VERSION : 0.1
   VAR
      MC_Interface : Array[0..12] of Struct
         Data_from_MC : Struct   // Signal from the mould carrier to the machine
            Automatic_mode : Bool;   // Mouldcarrier is in automatic mode and ready for production
            Selected : Bool;   // Mouldcarrier is selected
            Shot_preperation : Bool;   // Set shot preperation
            Shot_release : Bool;   // Set shot release
            Robot_release : Bool;   // Release move robot into MC
            Vacuum_on : Bool;   // Vacuum pump on from MC
            CP_forward : Bool;   // Cleaning piston forward from MC
            Com_control : Bool;   // Communication control
            Toolcode : Byte;   // Toolcode from MC
            Temperature_1 : Int;   // Temperature 1 from MC
            Temperature_2 : Int;   // Temperature 2 from MC
            Angle_frame_foaming_pos : Real;   // Angle (°) frame in foaming position
            Spare_10 : Word;
            Spare_12 : Word;
            Spare_14 : Word;
         END_STRUCT;
         Data_to_MC : Struct   // Signal from the machine to the mould carrier
            Automatic_mode : Bool;   // Foaming machine ready for production
            Service_mode : Bool;   // Shot simmulation active
            MH_selected : Bool;   // Mixinghead is selected
            Shot_runs : Bool;   // Shot runs
            Shot_end : Bool;   // Shot end
            Fault : Bool;   // Fault during shot
            Robot_out_of_MC : Bool;   // Robot out of mould carrier (to close the MC)
            Com_Control : Bool;   // Communication control
            Toolcode : Byte;   // Toolcode copy from foaming machine
            Spare_2 : Word;
            Spare_4 : Word;
            Spare_6 : Word;
            Spare_8 : Word;
            Spare_10 : Word;
            Spare_12 : Word;
            Spare_14 : Word;
         END_STRUCT;
      END_STRUCT;
   END_VAR
BEGIN
   MC_Interface[0].Data_to_MC.Spare_8 := 16#0000;
   MC_Interface[0].Data_to_MC.Spare_6 := 16#0000;
   MC_Interface[0].Data_to_MC.Spare_4 := 16#0000;
   MC_Interface[0].Data_to_MC.Spare_2 := 16#0000;
   MC_Interface[0].Data_to_MC.Toolcode := 16#00;
   MC_Interface[0].Data_to_MC.Com_Control := FALSE;
   MC_Interface[0].Data_to_MC.Robot_out_of_MC := FALSE;
   MC_Interface[0].Data_to_MC.Fault := FALSE;
   MC_Interface[0].Data_to_MC.Shot_end := FALSE;
   MC_Interface[0].Data_to_MC.Shot_runs := FALSE;
   MC_Interface[0].Data_to_MC.MH_selected := FALSE;
   MC_Interface[0].Data_to_MC.Service_mode := FALSE;
   MC_Interface[0].Data_to_MC.Automatic_mode := FALSE;
   MC_Interface[0].Data_from_MC.Automatic_mode := FALSE;
   MC_Interface[0].Data_from_MC.Selected := FALSE;
   MC_Interface[0].Data_from_MC.Shot_preperation := FALSE;
   MC_Interface[0].Data_from_MC.Shot_release := FALSE;
   MC_Interface[0].Data_from_MC.Robot_release := FALSE;
   MC_Interface[0].Data_from_MC.Vacuum_on := FALSE;
   MC_Interface[0].Data_from_MC.CP_forward := FALSE;
   MC_Interface[0].Data_from_MC.Com_control := FALSE;
   MC_Interface[0].Data_from_MC.Toolcode := 16#02;
   MC_Interface[0].Data_from_MC.Temperature_1 := 16#0000;
   MC_Interface[0].Data_from_MC.Temperature_2 := 16#0000;
   MC_Interface[0].Data_from_MC.Angle_frame_foaming_pos := 16#0000;
END_DATA_BLOCK

DATA_BLOCK "DB009_Faults"   // DB9
TITLE = State signals of fault handling
{ S7_Optimized_Access := 'FALSE' }
AUTHOR : KT242
VERSION : 0.1
   VAR
      Fault_State_Grp_1_M1 : Bool := FALSE;   // In der Steuerung wurde eine Störung der Gruppe 1 der Maschine 1 festgestellt
      Fault_State_Grp_2_M1 : Bool := FALSE;   // In der Steuerung wurde eine Störung der Gruppe 2 der Maschine 1 festgestellt
      Fault_State_Grp_3_M1 : Bool := FALSE;   // In der Steuerung wurde eine Störung der Gruppe 3 der Maschine 1 festgestellt
      Fault_State_Grp_1_M2 : Bool := FALSE;   // In der Steuerung wurde eine Störung der Gruppe 1 der Maschine 2 festgestellt
      Fault_State_Grp_2_M2 : Bool := FALSE;   // In der Steuerung wurde eine Störung der Gruppe 2 der Maschine 2 festgestellt
      Fault_State_Grp_3_M2 : Bool := FALSE;   // In der Steuerung wurde eine Störung der Gruppe 3 der Maschine 2 festgestellt
      Fault_State_Grp_1_M3 : Bool := FALSE;   // In der Steuerung wurde eine Störung der Gruppe 1 der Maschine 3 festgestellt
      Fault_State_Grp_2_M3 : Bool := FALSE;   // In der Steuerung wurde eine Störung der Gruppe 2 der Maschine 3 festgestellt
      Fault_State_Grp_3_M3 : Bool := FALSE;   // In der Steuerung wurde eine Störung der Gruppe 3 der Maschine 3 festgestellt
      Fault_State_Grp_1_M4 : Bool := FALSE;   // In der Steuerung wurde eine Störung der Gruppe 1 der Maschine 4 festgestellt
      Fault_State_Grp_2_M4 : Bool := FALSE;   // In der Steuerung wurde eine Störung der Gruppe 2 der Maschine 4 festgestellt
      Fault_State_Grp_3_M4 : Bool := FALSE;   // In der Steuerung wurde eine Störung der Gruppe 3 der Maschine 4 festgestellt
      Fault_State_Grp_1_ExtP : Bool := FALSE;   // In der Steuerung wurde eine Störung der Gruppe 1 der Fremdanlage festgestellt
      Fault_State_Grp_2_ExtP : Bool := FALSE;   // In der Steuerung wurde eine Störung der Gruppe 2 der Fremdanlage festgestellt
      Fault_State_Grp_3_ExtP : Bool := FALSE;   // In der Steuerung wurde eine Störung der Gruppe 3 der Fremdanlage festgestellt
      Fault_State_Grp_1_3_Exist : Bool := FALSE;   // In der Steuerung wurde eine Störung der Gruppe 1- 3 festgestellt
      Faultschanging_M1 : Bool := FALSE;   // Änderungsbit für die Signalauswertung // Hupe+ Lampe Maschine 1
      Faultschanging_M2 : Bool := FALSE;   // Änderungsbit für die Signalauswertung // Hupe+ Lampe Maschine 2
      Faultschanging_M3 : Bool := FALSE;   // Änderungsbit für die Signalauswertung // Hupe+ Lampe Maschine 3
      Faultschanging_M4 : Bool := FALSE;   // Änderungsbit für die Signalauswertung // Hupe+ Lampe Maschine 4
      Faultschanging_ExtP : Bool := FALSE;   // Änderungsbit für die Signalauswertung // Hupe+ Lampe Fremdanlage
      Reserve_2_5 : Bool := FALSE;
      Reserve_2_6 : Bool := FALSE;
      Reserve_2_7 : Bool := FALSE;
      HF_FaultsQuitOB35 : Bool := FALSE;   // Resetbit for faults in OB 35
      HF_Faults_Quit : Bool := FALSE;   // Flankenhilfsmerker für die Störungsquittierung
      HF_Horn : Bool := FALSE;   // Hilfsmerker für die Hupenansteuerung
      Faults_Reset_FKT_M1 : Bool := FALSE;   // Störungsbildung in den Funktionen der Maschine 1 zurücksetzen
      Faults_Reset_FKT_M2 : Bool := FALSE;   // Störungsbildung in den Funktionen der Maschine 2 zurücksetzen
      Faults_Reset_FKT_M3 : Bool := FALSE;   // Störungsbildung in den Funktionen der Maschine 3 zurücksetzen
      Faults_Reset_FKT_M4 : Bool := FALSE;   // Störungsbildung in den Funktionen der Maschine 4 zurücksetzen
      Faults_Reset_FKT_ExtP : Bool := FALSE;   // Störungsbildung in den Funktionen der Fremdanlage zurücksetzen
      Faults_Reset_Group : Bool := FALSE;   // Störungsbildung in den Störungsbausteinenzurücksetzen
      FaultPC_Level_1 : Bool := FALSE;
      FaultPC_Level_2 : Bool := FALSE;
      FaultPC_Level_3 : Bool := FALSE;
      Spare_6_3 : Bool := FALSE;
      Spare_6_4 : Bool := FALSE;
      Faults_FKT_Grp_1_M1 : Bool := FALSE;   // In der Steuerung wurde eine Störung der Gruppe 1 der Maschine 1 festgestellt
      Faults_FKT_Grp_2_M1 : Bool := FALSE;   // In der Steuerung wurde eine Störung der Gruppe 2 der Maschine 1 festgestellt
      Faults_FKT_Grp_3_M1 : Bool := FALSE;   // In der Steuerung wurde eine Störung der Gruppe 3 der Maschine 1 festgestellt
      Faults_FKT_Grp_1_M2 : Bool := FALSE;   // In der Steuerung wurde eine Störung der Gruppe 1 der Maschine 2 festgestellt
      Faults_FKT_Grp_2_M2 : Bool := FALSE;   // In der Steuerung wurde eine Störung der Gruppe 2 der Maschine 2 festgestellt
      Faults_FKT_Grp_3_M2 : Bool := FALSE;   // In der Steuerung wurde eine Störung der Gruppe 3 der Maschine 2 festgestellt
      Faults_FKT_Grp_1_M3 : Bool := FALSE;   // In der Steuerung wurde eine Störung der Gruppe 1 der Maschine 3 festgestellt
      Faults_FKT_Grp_2_M3 : Bool := FALSE;   // In der Steuerung wurde eine Störung der Gruppe 2 der Maschine 3 festgestellt
      Faults_FKT_Grp_3_M3 : Bool := FALSE;   // In der Steuerung wurde eine Störung der Gruppe 3 der Maschine 3 festgestellt
      Faults_FKT_Grp_1_M4 : Bool := FALSE;   // In der Steuerung wurde eine Störung der Gruppe 1 der Maschine 4 festgestellt
      Faults_FKT_Grp_2_M4 : Bool := FALSE;   // In der Steuerung wurde eine Störung der Gruppe 2 der Maschine 4 festgestellt
      Faults_FKT_Grp_3_M4 : Bool := FALSE;   // In der Steuerung wurde eine Störung der Gruppe 3 der Maschine 4 festgestellt
      Faults_FKT_Grp_1_ExtP : Bool := FALSE;   // In der Steuerung wurde eine Störung der Gruppe 1 der Fremdanlage festgestellt
      Faults_FKT_Grp_2_ExtP : Bool := FALSE;   // In der Steuerung wurde eine Störung der Gruppe 2 der Fremdanlage festgestellt
      Faults_FKT_Grp_3_ExtP : Bool := FALSE;   // In der Steuerung wurde eine Störung der Gruppe 3 der Fremdanlage festgestellt
      Spare_8_7 : Bool := FALSE;
      NewMessage_M1 : Bool := FALSE;   // New message comes up at machine 1
      NewMessage_M2 : Bool := FALSE;   // New message comes up at machine 2
      NewMessage_M3 : Bool := FALSE;   // New message comes up at machine 3
      NewMessage_M4 : Bool := FALSE;   // New message comes up at machine 4
      GoneMessage_M1 : Bool := TRUE;   // Message is no longer active machine 1
      GoneMessage_M2 : Bool := FALSE;   // Message is no longer active machine 2
      GoneMessage_M3 : Bool := FALSE;   // Message is no longer active machine 3
      GoneMessage_M4 : Bool := FALSE;   // Message is no longer active machine 4
      MessageChangedToVisu : Bool := TRUE;   // Signal to visualisation -> show fault messages and messages
      MessageChangedNext : Bool := TRUE;
      Spare_10_02 : Bool := FALSE;
      Spare_10_03 : Bool := FALSE;
      Spare_10_04 : Bool := FALSE;
      Spare_10_05 : Bool := FALSE;
      Spare_10_06 : Bool := FALSE;
      Spare_10_07 : Bool := FALSE;
   END_VAR
BEGIN
END_DATA_BLOCK

DATA_BLOCK "DB_MouldEditor_HMI"   // DB10
{ S7_Optimized_Access := 'FALSE' }
VERSION : 0.1
   VAR
      uData : "typeMouldEditor_HMI";   // Data for mould editor HMI
   END_VAR
BEGIN
END_DATA_BLOCK

DATA_BLOCK "FB_MouldEditor_HMI_DB"   // DB13
{ S7_Optimized_Access := 'FALSE' }
VERSION : 0.1
"FB_MouldEditor_HMI"
BEGIN
END_DATA_BLOCK

DATA_BLOCK "DB14_TP_Shortcuts"   // DB14
{ S7_Optimized_Access := 'TRUE' }
VERSION : 0.1
   VAR
      TP_Shortcuts : Struct
         ButtonNo : Struct
            "0" : Bool := FALSE;
            "1" : Bool := FALSE;
            "2" : Bool := FALSE;
            "3" : Bool := FALSE;
            "4" : Bool := FALSE;
            "5" : Bool := FALSE;
            "6" : Bool := FALSE;
            "7" : Bool := FALSE;
         END_STRUCT;
         PageNo : Struct
            "0" : Int := 0;
            "1" : Int := 0;
            "2" : Int := 15;
            "3" : Int := 0;
            "4" : Int := 9;
            "5" : Int := 0;
            "6" : Int := 100;
            "7" : Int := 9020;
         END_STRUCT;
         Page_active : Struct
            "0" : Bool := FALSE;
            "1" : Bool := FALSE;
            "2" : Bool := FALSE;
            "3" : Bool := FALSE;
            "4" : Bool := FALSE;
            "5" : Bool := FALSE;
            "6" : Bool := FALSE;
            "7" : Bool := FALSE;
         END_STRUCT;
      END_STRUCT;
   END_VAR
BEGIN
END_DATA_BLOCK

DATA_BLOCK "DB025_Oszilloskop"   // DB25
{ S7_Optimized_Access := 'FALSE' }
VERSION : 0.1
   VAR
      Graph : Array[1..10] of Struct
         Auswahl : Int;
         Nummer : Int;
         Komponente : Int;
         Sensor : Int;
         DB_Nummer : Word;
         Adresse : Int;
         Skalierung : Real;
         Wert : Real;
         Bit : Int;
      END_STRUCT;
      SkalierungGraphLinks : Struct
         Startwert : Int := 0;
         Ebdwert : Int := 200;
      END_STRUCT;
      SkalierungGraphRechts : Struct
         Startwert : Int := 0;
         Ebdwert : Int := 220;
      END_STRUCT;
   END_VAR
BEGIN
   Graph[1].Skalierung := 1.0;
   Graph[2].Skalierung := 1.0;
   Graph[3].Skalierung := 1.0;
   Graph[4].Skalierung := 1.0;
   Graph[5].Skalierung := 1.0;
   Graph[6].Skalierung := 1.0;
   Graph[7].Skalierung := 1.0;
   Graph[8].Skalierung := 1.0;
   Graph[9].Skalierung := 1.0;
   Graph[10].Skalierung := 1.0;
   Graph[1].Auswahl := 30;
   Graph[1].Nummer := 0;
   Graph[1].Komponente := 1;
   Graph[1].Sensor := 1;
   Graph[1].DB_Nummer := 16#0000;
   Graph[1].Adresse := 0;
   Graph[1].Wert := 0.0;
   Graph[1].Bit := 0;
   Graph[2].Auswahl := 30;
   Graph[2].Nummer := 1;
   Graph[2].Komponente := 2;
   Graph[2].Sensor := 1;
   Graph[2].DB_Nummer := 16#0000;
   Graph[2].Adresse := 0;
   Graph[2].Wert := 0.0;
   Graph[2].Bit := 0;
   Graph[3].Auswahl := 0;
   Graph[3].Nummer := 0;
   Graph[3].Komponente := 0;
   Graph[3].Sensor := 0;
   Graph[3].DB_Nummer := 16#0000;
   Graph[3].Adresse := 0;
   Graph[3].Wert := 0.0;
   Graph[3].Bit := 0;
   Graph[4].Auswahl := 0;
   Graph[4].Nummer := 0;
   Graph[4].Komponente := 0;
   Graph[4].Sensor := 0;
   Graph[4].DB_Nummer := 16#0000;
   Graph[4].Adresse := 0;
   Graph[4].Wert := 0.0;
   Graph[4].Bit := 0;
   Graph[5].Auswahl := 0;
   Graph[5].Nummer := 0;
   Graph[5].Komponente := 0;
   Graph[5].Sensor := 0;
   Graph[5].DB_Nummer := 16#0000;
   Graph[5].Adresse := 0;
   Graph[5].Wert := 0.0;
   Graph[5].Bit := 0;
   Graph[6].Auswahl := 0;
   Graph[6].Nummer := 0;
   Graph[6].Komponente := 0;
   Graph[6].Sensor := 0;
   Graph[6].DB_Nummer := 16#0000;
   Graph[6].Adresse := 0;
   Graph[6].Wert := 0.0;
   Graph[6].Bit := 0;
   Graph[7].Auswahl := 20;
   Graph[7].Nummer := 1;
   Graph[7].Komponente := 1;
   Graph[7].Sensor := 2;
   Graph[7].DB_Nummer := 16#0000;
   Graph[7].Adresse := 0;
   Graph[7].Wert := 1.8;
   Graph[7].Bit := 0;
   Graph[8].Auswahl := 20;
   Graph[8].Nummer := 1;
   Graph[8].Komponente := 2;
   Graph[8].Sensor := 2;
   Graph[8].DB_Nummer := 16#0000;
   Graph[8].Adresse := 0;
   Graph[8].Wert := 2.2;
   Graph[8].Bit := 0;
   Graph[9].Auswahl := 0;
   Graph[9].Nummer := 0;
   Graph[9].Komponente := 0;
   Graph[9].Sensor := 0;
   Graph[9].DB_Nummer := 16#0000;
   Graph[9].Adresse := 0;
   Graph[9].Wert := 0.0;
   Graph[9].Bit := 0;
   Graph[10].Auswahl := 0;
   Graph[10].Nummer := 0;
   Graph[10].Komponente := 0;
   Graph[10].Sensor := 0;
   Graph[10].DB_Nummer := 16#0000;
   Graph[10].Adresse := 0;
   Graph[10].Wert := 0.0;
   Graph[10].Bit := 0;
END_DATA_BLOCK

DATA_BLOCK "BalluffReader_1"   // DB30
{ S7_Optimized_Access := 'FALSE' }
AUTHOR : Serrano
FAMILY : Ident
NAME : BIS60X2
VERSION : 1.8
"FB030_BallufReader"
BEGIN
END_DATA_BLOCK

DATA_BLOCK "BalluffReader_2"   // DB31
{ S7_Optimized_Access := 'FALSE' }
AUTHOR : Serrano
FAMILY : Ident
NAME : BIS60X2
VERSION : 1.8
"FB030_BallufReader"
BEGIN
END_DATA_BLOCK

DATA_BLOCK "BalluffReader"   // DB32
{ S7_Optimized_Access := 'FALSE' }
VERSION : 0.1
   VAR
      ReadWriteHead1 : Struct
         Command_Write : Bool := FALSE;
         FHM_Command_Write : Bool := FALSE;
         HM_Command_Write : Bool := FALSE;
         Command_Read : Bool := FALSE;
         FHM_Command_Read : Bool := FALSE;
         HM_Command_Read : Bool := FALSE;
         FHM_Read_Auto : Bool := FALSE;   // FHM Automatisch Lesen nach Schreiben
         HM_Read_Auto : Bool := FALSE;   // HM Automatisch Lesen nach Schreiben
         FHM_Code_was_readed : Bool := FALSE;   // FHM Code gelesen
         HM_Code_was_readed : Bool := FALSE;   // HM Code gelesen
         Code_was_readed : Bool := FALSE;   // HM Code gelesen
         FHM_Writing_was_activ : Bool := FALSE;   // FHM Beschreiben Datenträger war aktiv
         HM_Writing_was_activ : Bool := FALSE;   // HM Beschreiben Datenträger war aktiv
         FHM_Start_Zyklus : Bool;
         Spare_1_6 : Bool;
         Spare_1_7 : Bool;
         Fault_01 : Bool := FALSE;   // Kein Datenträger vorhanden
         Fault_02 : Bool := FALSE;   // Fehler beim Lesen
         Fault_03 : Bool := FALSE;   // Lesen abgebrochen, da Datenträger entfernt wurde
         Fault_04 : Bool := FALSE;   // Fehler beim Schreiben
         Fault_05 : Bool := FALSE;   // Schreiben abgebrochen, da Datenträger entfernt wurde
         Fault_06 : Bool := FALSE;   // Zugriffsfehler auf Speicher
         Fault_07 : Bool := FALSE;   // Falsche Befehlskennung oder Anzahl Byte bei einem Schreib-/Lesebefehl ist 0
         Fault_08 : Bool := FALSE;   // Kabelbruch des angewählten Schreib-/Lesekopfs
         Fault_09 : Bool := FALSE;   // EEProm in der Auswerteeinheit defekt
         Fault_10 : Bool := FALSE;   // Kommunikation zum Datenträger gestört
         Fault_11 : Bool := FALSE;   // Inhalt der 1. und 2. Bitleiste sind ungleich
         Fault_12 : Bool := FALSE;   // Startadresse + Anzahl Bytes > Speicherbereich in Initialisierung angegeben
         Fault_13 : Bool := FALSE;   // Ungültige max. Anzahl Schreibzyklen in Initialisierung angegeben
         Fault_14 : Bool := FALSE;   // max. Anzahl von 1kByte in Initialisierung überschritten
         Fault_15 : Bool := FALSE;   // Überwachung der Initialisierung bringt keine Übereinstimmung.
         Fault_16 : Bool := FALSE;   // Datenträger nicht initialisiert. Alle Bytes noch 00h
         Spare_4 : Byte;
         Spare_5 : Byte;
         Spare_6 : Byte;
         Spare_7 : Byte;
         TM_RFID : S5Time := S5T#4s;   // Überwachungszeit zum lesen/schreiben
         Send : Struct
            Program : Int;
            Text : Array[1..30] of Char;
         END_STRUCT;
         Receive : Struct
            Program : Int;
            Text : Array[1..30] of Char;
         END_STRUCT;
      END_STRUCT;
      ReadWriteHead2 : Struct
         Command_Write : Bool := FALSE;
         FHM_Command_Write : Bool := FALSE;
         HM_Command_Write : Bool := FALSE;
         Command_Read : Bool := FALSE;
         FHM_Command_Read : Bool := FALSE;
         HM_Command_Read : Bool := FALSE;
         FHM_Read_Auto : Bool := FALSE;   // FHM Automatisch Lesen nach Schreiben
         HM_Read_Auto : Bool := FALSE;   // HM Automatisch Lesen nach Schreiben
         FHM_Code_was_readed : Bool := FALSE;   // FHM Code gelesen
         HM_Code_was_readed : Bool := FALSE;   // HM Code gelesen
         Code_was_readed : Bool := FALSE;   // HM Code gelesen für Zylinder zurück
         FHM_Writing_was_activ : Bool := FALSE;   // FHM Beschreiben Datenträger war aktiv
         HM_Writing_was_activ : Bool := FALSE;   // HM Beschreiben Datenträger war aktiv
         FHM_Start_Zyklus : Bool;
         Spare_1_6 : Bool;
         Spare_1_7 : Bool;
         Fault_01 : Bool := FALSE;   // Kein Datenträger vorhanden
         Fault_02 : Bool := FALSE;   // Fehler beim Lesen
         Fault_03 : Bool := FALSE;   // Lesen abgebrochen, da Datenträger entfernt wurde
         Fault_04 : Bool := FALSE;   // Fehler beim Schreiben
         Fault_05 : Bool := FALSE;   // Schreiben abgebrochen, da Datenträger entfernt wurde
         Fault_06 : Bool := FALSE;   // Zugriffsfehler auf Speicher
         Fault_07 : Bool := FALSE;   // Falsche Befehlskennung oder Anzahl Byte bei einem Schreib-/Lesebefehl ist 0
         Fault_08 : Bool := FALSE;   // Kabelbruch des angewählten Schreib-/Lesekopfs
         Fault_09 : Bool := FALSE;   // EEProm in der Auswerteeinheit defekt
         Fault_10 : Bool := FALSE;   // Kommunikation zum Datenträger gestört
         Fault_11 : Bool := FALSE;   // Inhalt der 1. und 2. Bitleiste sind ungleich
         Fault_12 : Bool := FALSE;   // Startadresse + Anzahl Bytes > Speicherbereich in Initialisierung angegeben
         Fault_13 : Bool := FALSE;   // Ungültige max. Anzahl Schreibzyklen in Initialisierung angegeben
         Fault_14 : Bool := FALSE;   // max. Anzahl von 1kByte in Initialisierung überschritten
         Fault_15 : Bool := FALSE;   // Überwachung der Initialisierung bringt keine Übereinstimmung.
         Fault_16 : Bool := FALSE;   // Datenträger nicht initialisiert. Alle Bytes noch 00h
         Spare_4 : Byte;
         Spare_5 : Byte;
         Spare_6 : Byte;
         Spare_7 : Byte;
         TM_RFID : S5Time := S5T#4s;   // Überwachungszeit zum lesen/schreiben
         Send : Struct
            Program : Int;
            Text : Array[1..30] of Char;
         END_STRUCT;
         Receive : Struct
            Program : Int;
            Text : Array[1..30] of Char;
         END_STRUCT;
      END_STRUCT;
   END_VAR
BEGIN
END_DATA_BLOCK

DATA_BLOCK "DB110_Interf_Program_M1"   // DB110
TITLE = Signal between pouring machine and external plant parts
{ S7_Optimized_Access := 'FALSE' }
AUTHOR : KT242
VERSION : 0.1
   VAR
      Bits : Struct
         Ageflag : Bool := TRUE;
         Stop_Cycle : Bool := FALSE;
         startbutton_activated : Bool := FALSE;
         HF_StopCycleWHileToolDisabled : Bool := FALSE;
         F_StopCycleWHileToolDisabled : Bool := FALSE;
         LastShotAtThisMachine : Bool := FALSE;
         PulseShotEnd : Bool := FALSE;
         PulseToolFinished : Bool := FALSE;
         HF_FP_PulseToolFinished : Bool := TRUE;
         LockAutoCycleStart : Bool := FALSE;
         MouldNotReleased : Bool := FALSE;
         HF_FP_MouldNotReleased : Bool := FALSE;
         LastStandbyTimeTool : Bool := FALSE;
         PulseCycleEnd : Bool := FALSE;
         HF_FP_CycleNotRunning : Bool := TRUE;
         HF_FP_ResetProgramNo : Bool := FALSE;
      END_STRUCT;
      Putin_FIFOlist : "UDT001_DWord_1_32";
      FIRST : Int := 0;
      SECOND : Int := 0;
      FIFO : Struct
         FIFO_01 : Word := 16#0000;
         FIFO_02 : Word := 16#0000;
         FIFO_03 : Word := 16#0000;
         FIFO_04 : Word := 16#0000;
         FIFO_05 : Word := 16#0000;
         FIFO_06 : Word := 16#0000;
         FIFO_07 : Word := 16#0000;
         FIFO_08 : Word := 16#0000;
         FIFO_09 : Word := 16#0000;
         FIFO_10 : Word := 16#0000;
         FIFO_11 : Word := 16#0000;
         FIFO_12 : Word := 16#0000;
         FIFO_13 : Word := 16#0000;
         FIFO_14 : Word := 16#0000;
         FIFO_15 : Word := 16#0000;
         FIFO_16 : Word := 16#0000;
         FIFO_17 : Word := 16#0000;
         FIFO_18 : Word := 16#0000;
         FIFO_19 : Word := 16#0000;
         FIFO_20 : Word := 16#0000;
         FIFO_21 : Word := 16#0000;
         FIFO_22 : Word := 16#0000;
         FIFO_23 : Word := 16#0000;
         FIFO_24 : Word := 16#0000;
         FIFO_25 : Word := 16#0000;
         FIFO_26 : Word := 16#0000;
         FIFO_27 : Word := 16#0000;
         FIFO_28 : Word := 16#0000;
         FIFO_29 : Word := 16#0000;
         FIFO_30 : Word := 16#0000;
         FIFO_31 : Word := 16#0000;
         FIFO_32 : Word := 16#0000;
      END_STRUCT;
      Test_M01 : "UDT115_Test";
      Test_M02 : "UDT115_Test";
      Test_M03 : "UDT115_Test";
      Test_M04 : "UDT115_Test";
      Status_IF : Array[1..16] of "UDT112_IF_UP_MC";
      HM_MC_Fault : "UDT001_DWord_1_32";
      HM_MC_Shotend : "UDT001_DWord_1_32";
      HM_MC_Lamp : "UDT001_DWord_1_32";
      HM_MC_mould_Closing : "UDT001_DWord_1_32";
      HM_MC_spare : "UDT001_DWord_1_32";
      Program_is_active : "UDT001_DWord_1_32";
      Program_No_01 : Word := 16#0000;
      Program_No_02 : Word := 16#0000;
      Program_No_03 : Word := 16#0000;
      Program_No_04 : Word := 16#0000;
      Program_No_05 : Word := 16#0000;
      Program_No_06 : Word := 16#0000;
      Program_No_07 : Word := 16#0000;
      Program_No_08 : Word := 16#0000;
      Robot_01 : "ABB_IRC5_Status";
      Mixingheadcleaner_01 : "UDT118_MH_Cleaner";
      Bandfilter_01 : "UDT119_Bandfilter";
      Robot_02 : "ABB_IRC5_Status";
      Mixingheadcleaner_02 : "UDT118_MH_Cleaner";
      Bandfilter_02 : "UDT119_Bandfilter";
      MixingHeadNo : Int := 0;
      Signals_ExPlant : Array[1..4] of "UDT1114_IF_Signals";
      Status_ExPlant : Array[1..4] of "UDT114_IF_externalPlant";
   END_VAR
BEGIN
   Putin_FIFOlist."25" := FALSE;
   Putin_FIFOlist."26" := FALSE;
   Putin_FIFOlist."27" := FALSE;
   Putin_FIFOlist."28" := FALSE;
   Putin_FIFOlist."29" := FALSE;
   Putin_FIFOlist."30" := FALSE;
   Putin_FIFOlist."31" := FALSE;
   Putin_FIFOlist."32" := FALSE;
   Putin_FIFOlist."17" := FALSE;
   Putin_FIFOlist."18" := FALSE;
   Putin_FIFOlist."19" := FALSE;
   Putin_FIFOlist."20" := FALSE;
   Putin_FIFOlist."21" := FALSE;
   Putin_FIFOlist."22" := FALSE;
   Putin_FIFOlist."23" := FALSE;
   Putin_FIFOlist."24" := FALSE;
   Putin_FIFOlist."09" := FALSE;
   Putin_FIFOlist."10" := FALSE;
   Putin_FIFOlist."11" := FALSE;
   Putin_FIFOlist."12" := FALSE;
   Putin_FIFOlist."13" := FALSE;
   Putin_FIFOlist."14" := FALSE;
   Putin_FIFOlist."15" := FALSE;
   Putin_FIFOlist."16" := FALSE;
   Putin_FIFOlist."01" := FALSE;
   Putin_FIFOlist."02" := FALSE;
   Putin_FIFOlist."03" := FALSE;
   Putin_FIFOlist."04" := FALSE;
   Putin_FIFOlist."05" := FALSE;
   Putin_FIFOlist."06" := FALSE;
   Putin_FIFOlist."07" := FALSE;
   Putin_FIFOlist."08" := FALSE;
   Test_M01.Test_runs := FALSE;
   Test_M01.Test_K1 := FALSE;
   Test_M01.Test_K2 := FALSE;
   Test_M01.Test_K3 := FALSE;
   Test_M01.Test_K4 := FALSE;
   Test_M01.Start_to_Cycle := FALSE;
   Test_M01.Stop_to_Cycle := FALSE;
   Test_M01.Spare_0_7 := FALSE;
   Test_M01.Spare_Byte := 16#00;
   Test_M02.Test_runs := FALSE;
   Test_M02.Test_K1 := FALSE;
   Test_M02.Test_K2 := FALSE;
   Test_M02.Test_K3 := FALSE;
   Test_M02.Test_K4 := FALSE;
   Test_M02.Start_to_Cycle := FALSE;
   Test_M02.Stop_to_Cycle := FALSE;
   Test_M02.Spare_0_7 := FALSE;
   Test_M02.Spare_Byte := 16#00;
   Test_M03.Test_runs := FALSE;
   Test_M03.Test_K1 := FALSE;
   Test_M03.Test_K2 := FALSE;
   Test_M03.Test_K3 := FALSE;
   Test_M03.Test_K4 := FALSE;
   Test_M03.Start_to_Cycle := FALSE;
   Test_M03.Stop_to_Cycle := FALSE;
   Test_M03.Spare_0_7 := FALSE;
   Test_M03.Spare_Byte := 16#00;
   Test_M04.Test_runs := FALSE;
   Test_M04.Test_K1 := FALSE;
   Test_M04.Test_K2 := FALSE;
   Test_M04.Test_K3 := FALSE;
   Test_M04.Test_K4 := FALSE;
   Test_M04.Start_to_Cycle := FALSE;
   Test_M04.Stop_to_Cycle := FALSE;
   Test_M04.Spare_0_7 := FALSE;
   Test_M04.Spare_Byte := 16#00;
   HM_MC_Fault."25" := FALSE;
   HM_MC_Fault."26" := FALSE;
   HM_MC_Fault."27" := FALSE;
   HM_MC_Fault."28" := FALSE;
   HM_MC_Fault."29" := FALSE;
   HM_MC_Fault."30" := FALSE;
   HM_MC_Fault."31" := FALSE;
   HM_MC_Fault."32" := FALSE;
   HM_MC_Fault."17" := FALSE;
   HM_MC_Fault."18" := FALSE;
   HM_MC_Fault."19" := FALSE;
   HM_MC_Fault."20" := FALSE;
   HM_MC_Fault."21" := FALSE;
   HM_MC_Fault."22" := FALSE;
   HM_MC_Fault."23" := FALSE;
   HM_MC_Fault."24" := FALSE;
   HM_MC_Fault."09" := FALSE;
   HM_MC_Fault."10" := FALSE;
   HM_MC_Fault."11" := FALSE;
   HM_MC_Fault."12" := FALSE;
   HM_MC_Fault."13" := FALSE;
   HM_MC_Fault."14" := FALSE;
   HM_MC_Fault."15" := FALSE;
   HM_MC_Fault."16" := FALSE;
   HM_MC_Fault."01" := FALSE;
   HM_MC_Fault."02" := FALSE;
   HM_MC_Fault."03" := FALSE;
   HM_MC_Fault."04" := FALSE;
   HM_MC_Fault."05" := FALSE;
   HM_MC_Fault."06" := FALSE;
   HM_MC_Fault."07" := FALSE;
   HM_MC_Fault."08" := FALSE;
   HM_MC_Shotend."25" := FALSE;
   HM_MC_Shotend."26" := FALSE;
   HM_MC_Shotend."27" := FALSE;
   HM_MC_Shotend."28" := FALSE;
   HM_MC_Shotend."29" := FALSE;
   HM_MC_Shotend."30" := FALSE;
   HM_MC_Shotend."31" := FALSE;
   HM_MC_Shotend."32" := FALSE;
   HM_MC_Shotend."17" := FALSE;
   HM_MC_Shotend."18" := FALSE;
   HM_MC_Shotend."19" := FALSE;
   HM_MC_Shotend."20" := FALSE;
   HM_MC_Shotend."21" := FALSE;
   HM_MC_Shotend."22" := FALSE;
   HM_MC_Shotend."23" := FALSE;
   HM_MC_Shotend."24" := FALSE;
   HM_MC_Shotend."09" := FALSE;
   HM_MC_Shotend."10" := FALSE;
   HM_MC_Shotend."11" := FALSE;
   HM_MC_Shotend."12" := FALSE;
   HM_MC_Shotend."13" := FALSE;
   HM_MC_Shotend."14" := FALSE;
   HM_MC_Shotend."15" := FALSE;
   HM_MC_Shotend."16" := FALSE;
   HM_MC_Shotend."01" := FALSE;
   HM_MC_Shotend."02" := FALSE;
   HM_MC_Shotend."03" := FALSE;
   HM_MC_Shotend."04" := FALSE;
   HM_MC_Shotend."05" := FALSE;
   HM_MC_Shotend."06" := FALSE;
   HM_MC_Shotend."07" := FALSE;
   HM_MC_Shotend."08" := FALSE;
   HM_MC_Lamp."25" := FALSE;
   HM_MC_Lamp."26" := FALSE;
   HM_MC_Lamp."27" := FALSE;
   HM_MC_Lamp."28" := FALSE;
   HM_MC_Lamp."29" := FALSE;
   HM_MC_Lamp."30" := FALSE;
   HM_MC_Lamp."31" := FALSE;
   HM_MC_Lamp."32" := FALSE;
   HM_MC_Lamp."17" := FALSE;
   HM_MC_Lamp."18" := FALSE;
   HM_MC_Lamp."19" := FALSE;
   HM_MC_Lamp."20" := FALSE;
   HM_MC_Lamp."21" := FALSE;
   HM_MC_Lamp."22" := FALSE;
   HM_MC_Lamp."23" := FALSE;
   HM_MC_Lamp."24" := FALSE;
   HM_MC_Lamp."09" := FALSE;
   HM_MC_Lamp."10" := FALSE;
   HM_MC_Lamp."11" := FALSE;
   HM_MC_Lamp."12" := FALSE;
   HM_MC_Lamp."13" := FALSE;
   HM_MC_Lamp."14" := FALSE;
   HM_MC_Lamp."15" := FALSE;
   HM_MC_Lamp."16" := FALSE;
   HM_MC_Lamp."01" := FALSE;
   HM_MC_Lamp."02" := FALSE;
   HM_MC_Lamp."03" := FALSE;
   HM_MC_Lamp."04" := FALSE;
   HM_MC_Lamp."05" := FALSE;
   HM_MC_Lamp."06" := FALSE;
   HM_MC_Lamp."07" := FALSE;
   HM_MC_Lamp."08" := FALSE;
   HM_MC_mould_Closing."25" := FALSE;
   HM_MC_mould_Closing."26" := FALSE;
   HM_MC_mould_Closing."27" := FALSE;
   HM_MC_mould_Closing."28" := FALSE;
   HM_MC_mould_Closing."29" := FALSE;
   HM_MC_mould_Closing."30" := FALSE;
   HM_MC_mould_Closing."31" := FALSE;
   HM_MC_mould_Closing."32" := FALSE;
   HM_MC_mould_Closing."17" := FALSE;
   HM_MC_mould_Closing."18" := FALSE;
   HM_MC_mould_Closing."19" := FALSE;
   HM_MC_mould_Closing."20" := FALSE;
   HM_MC_mould_Closing."21" := FALSE;
   HM_MC_mould_Closing."22" := FALSE;
   HM_MC_mould_Closing."23" := FALSE;
   HM_MC_mould_Closing."24" := FALSE;
   HM_MC_mould_Closing."09" := FALSE;
   HM_MC_mould_Closing."10" := FALSE;
   HM_MC_mould_Closing."11" := FALSE;
   HM_MC_mould_Closing."12" := FALSE;
   HM_MC_mould_Closing."13" := FALSE;
   HM_MC_mould_Closing."14" := FALSE;
   HM_MC_mould_Closing."15" := FALSE;
   HM_MC_mould_Closing."16" := FALSE;
   HM_MC_mould_Closing."01" := FALSE;
   HM_MC_mould_Closing."02" := FALSE;
   HM_MC_mould_Closing."03" := FALSE;
   HM_MC_mould_Closing."04" := FALSE;
   HM_MC_mould_Closing."05" := FALSE;
   HM_MC_mould_Closing."06" := FALSE;
   HM_MC_mould_Closing."07" := FALSE;
   HM_MC_mould_Closing."08" := FALSE;
   HM_MC_spare."25" := FALSE;
   HM_MC_spare."26" := FALSE;
   HM_MC_spare."27" := FALSE;
   HM_MC_spare."28" := FALSE;
   // 962 more start values not shown
END_DATA_BLOCK

DATA_BLOCK "DB119_Interface_Visu"   // DB119
TITLE = Signal between pouring machine and external plant parts
{ S7_Optimized_Access := 'FALSE' }
AUTHOR : KT242
VERSION : 0.1
   VAR
      "Inv.PrgNr" : Bool := TRUE;
      Profibus : Bool := FALSE;
      Paritätsbit : Bool := FALSE;
      ReadWriteDeviceNo : Int := 0;
      CopyDeviceNO : Int := 0;
      Read : Bool := FALSE;
      Write : Bool := FALSE;
      Copy : Bool := FALSE;
      Activ : Bool := FALSE;
      MouldCarrer : Array[0..12] of "UDT1111_MouldCarrier";
      APInterface : Array[0..12] of "UDT1112_APInterface";
   END_VAR
BEGIN
   APInterface[0].PrgNo := 16#FF;
   APInterface[0].ExtP_OK := TRUE;
   APInterface[0].Strobe := TRUE;
   APInterface[0].StrobeInv := TRUE;
   APInterface[0].MH_open := TRUE;
   APInterface[0].CP_forward := TRUE;
   APInterface[0].Preparation := TRUE;
   APInterface[0].Start_Cleaning := TRUE;
   APInterface[0].Stop := TRUE;
   APInterface[0].PU_OK := TRUE;
   APInterface[0].Strobe_quitt := TRUE;
   APInterface[0].cycle_run := TRUE;
   APInterface[0].ready_for_shot := TRUE;
   APInterface[0].shot_run := TRUE;
   APInterface[0].shot_end := TRUE;
   APInterface[0].Service_mode := TRUE;
   APInterface[0].CP_is_forward := TRUE;
   APInterface[0].Cleaning_finished := TRUE;
   APInterface[0].Reserve31 := TRUE;
   MouldCarrer[0].Preparation := FALSE;
   MouldCarrer[0].StartFoaming := FALSE;
   MouldCarrer[0].IN_Spare_01 := FALSE;
   MouldCarrer[0].IN_Spare_02 := FALSE;
   MouldCarrer[0].IN_Spare_03 := FALSE;
   MouldCarrer[0].IN_Spare_04 := FALSE;
   MouldCarrer[0].IN_Spare_05 := FALSE;
   MouldCarrer[0].IN_Spare_06 := FALSE;
   MouldCarrer[0].ShotEnds := FALSE;
   MouldCarrer[0].Break := FALSE;
   MouldCarrer[0].OUT_Spare_01 := FALSE;
   MouldCarrer[0].OUT_Spare_02 := FALSE;
   MouldCarrer[0].OUT_Spare_03 := FALSE;
   MouldCarrer[0].OUT_Spare_04 := FALSE;
   MouldCarrer[0].OUT_Spare_05 := FALSE;
   MouldCarrer[0].OUT_Spare_06 := FALSE;
   MouldCarrer[0].NoFault := FALSE;
   MouldCarrer[0].MachineAutomatic := FALSE;
   MouldCarrer[0].MHAutomatic := FALSE;
   MouldCarrer[0].RobotAutomatic := FALSE;
   MouldCarrer[0].WetShot := FALSE;
   MouldCarrer[0].CycleRun := FALSE;
   MouldCarrer[0].ReadyForShot := FALSE;
   MouldCarrer[0].ShotRun := FALSE;
   MouldCarrer[0].CPsisForward := FALSE;
   MouldCarrer[0].Status_Spare_01 := FALSE;
   MouldCarrer[0].Status_Spare_02 := FALSE;
   MouldCarrer[0].Status_Spare_03 := FALSE;
   MouldCarrer[0].Status_Spare_04 := FALSE;
   MouldCarrer[0].Status_Spare_05 := FALSE;
   MouldCarrer[0].Status_Spare_06 := FALSE;
   MouldCarrer[0].Status_Spare_07 := FALSE;
   MouldCarrer[0].ProgNumber := FALSE;
   MouldCarrer[0].Fault_01 := FALSE;
   MouldCarrer[0].Fault_02 := FALSE;
   MouldCarrer[0].Fault_03 := FALSE;
   MouldCarrer[0].Fault_04 := FALSE;
   MouldCarrer[0].Fault_05 := FALSE;
   MouldCarrer[0].Fault_06 := FALSE;
   MouldCarrer[0].Fault_07 := FALSE;
   MouldCarrer[0].Fault_08 := FALSE;
   MouldCarrer[1].Preparation := FALSE;
   MouldCarrer[1].StartFoaming := FALSE;
   MouldCarrer[1].IN_Spare_01 := FALSE;
   MouldCarrer[1].IN_Spare_02 := FALSE;
   MouldCarrer[1].IN_Spare_03 := FALSE;
   MouldCarrer[1].IN_Spare_04 := FALSE;
   MouldCarrer[1].IN_Spare_05 := FALSE;
   MouldCarrer[1].IN_Spare_06 := FALSE;
   MouldCarrer[1].ShotEnds := FALSE;
   MouldCarrer[1].Break := FALSE;
   MouldCarrer[1].OUT_Spare_01 := FALSE;
   MouldCarrer[1].OUT_Spare_02 := FALSE;
   MouldCarrer[1].OUT_Spare_03 := FALSE;
   MouldCarrer[1].OUT_Spare_04 := FALSE;
   MouldCarrer[1].OUT_Spare_05 := FALSE;
   MouldCarrer[1].OUT_Spare_06 := FALSE;
   MouldCarrer[1].NoFault := FALSE;
   MouldCarrer[1].MachineAutomatic := FALSE;
   MouldCarrer[1].MHAutomatic := FALSE;
   MouldCarrer[1].RobotAutomatic := FALSE;
   MouldCarrer[1].WetShot := FALSE;
   MouldCarrer[1].CycleRun := FALSE;
   MouldCarrer[1].ReadyForShot := FALSE;
   MouldCarrer[1].ShotRun := FALSE;
   MouldCarrer[1].CPsisForward := FALSE;
   MouldCarrer[1].Status_Spare_01 := FALSE;
   MouldCarrer[1].Status_Spare_02 := FALSE;
   MouldCarrer[1].Status_Spare_03 := FALSE;
   MouldCarrer[1].Status_Spare_04 := FALSE;
   MouldCarrer[1].Status_Spare_05 := FALSE;
   MouldCarrer[1].Status_Spare_06 := FALSE;
   MouldCarrer[1].Status_Spare_07 := FALSE;
   MouldCarrer[1].ProgNumber := FALSE;
   MouldCarrer[1].Fault_01 := FALSE;
   MouldCarrer[1].Fault_02 := FALSE;
   MouldCarrer[1].Fault_03 := FALSE;
   MouldCarrer[1].Fault_04 := FALSE;
   MouldCarrer[1].Fault_05 := FALSE;
   MouldCarrer[1].Fault_06 := FALSE;
   MouldCarrer[1].Fault_07 := FALSE;
   MouldCarrer[1].Fault_08 := FALSE;
   MouldCarrer[2].Preparation := FALSE;
   MouldCarrer[2].StartFoaming := FALSE;
   MouldCarrer[2].IN_Spare_01 := FALSE;
   MouldCarrer[2].IN_Spare_02 := FALSE;
   MouldCarrer[2].IN_Spare_03 := FALSE;
   MouldCarrer[2].IN_Spare_04 := FALSE;
   MouldCarrer[2].IN_Spare_05 := FALSE;
   MouldCarrer[2].IN_Spare_06 := FALSE;
   MouldCarrer[2].ShotEnds := FALSE;
   MouldCarrer[2].Break := FALSE;
   MouldCarrer[2].OUT_Spare_01 := FALSE;
   MouldCarrer[2].OUT_Spare_02 := FALSE;
   MouldCarrer[2].OUT_Spare_03 := FALSE;
   MouldCarrer[2].OUT_Spare_04 := FALSE;
   MouldCarrer[2].OUT_Spare_05 := FALSE;
   MouldCarrer[2].OUT_Spare_06 := FALSE;
   MouldCarrer[2].NoFault := FALSE;
   MouldCarrer[2].MachineAutomatic := FALSE;
   MouldCarrer[2].MHAutomatic := FALSE;
   MouldCarrer[2].RobotAutomatic := FALSE;
   MouldCarrer[2].WetShot := FALSE;
   MouldCarrer[2].CycleRun := FALSE;
   MouldCarrer[2].ReadyForShot := FALSE;
   MouldCarrer[2].ShotRun := FALSE;
   MouldCarrer[2].CPsisForward := FALSE;
   MouldCarrer[2].Status_Spare_01 := FALSE;
   MouldCarrer[2].Status_Spare_02 := FALSE;
   MouldCarrer[2].Status_Spare_03 := FALSE;
   MouldCarrer[2].Status_Spare_04 := FALSE;
   MouldCarrer[2].Status_Spare_05 := FALSE;
   MouldCarrer[2].Status_Spare_06 := FALSE;
   MouldCarrer[2].Status_Spare_07 := FALSE;
   MouldCarrer[2].ProgNumber := FALSE;
   MouldCarrer[2].Fault_01 := FALSE;
   MouldCarrer[2].Fault_02 := FALSE;
   MouldCarrer[2].Fault_03 := FALSE;
   MouldCarrer[2].Fault_04 := FALSE;
   MouldCarrer[2].Fault_05 := FALSE;
   MouldCarrer[2].Fault_06 := FALSE;
   MouldCarrer[2].Fault_07 := FALSE;
   MouldCarrer[2].Fault_08 := FALSE;
   MouldCarrer[3].Preparation := FALSE;
   MouldCarrer[3].StartFoaming := FALSE;
   MouldCarrer[3].IN_Spare_01 := FALSE;
   MouldCarrer[3].IN_Spare_02 := FALSE;
   MouldCarrer[3].IN_Spare_03 := FALSE;
   MouldCarrer[3].IN_Spare_04 := FALSE;
   MouldCarrer[3].IN_Spare_05 := FALSE;
   MouldCarrer[3].IN_Spare_06 := FALSE;
   MouldCarrer[3].ShotEnds := FALSE;
   MouldCarrer[3].Break := FALSE;
   MouldCarrer[3].OUT_Spare_01 := FALSE;
   MouldCarrer[3].OUT_Spare_02 := FALSE;
   MouldCarrer[3].OUT_Spare_03 := FALSE;
   MouldCarrer[3].OUT_Spare_04 := FALSE;
   MouldCarrer[3].OUT_Spare_05 := FALSE;
   MouldCarrer[3].OUT_Spare_06 := FALSE;
   MouldCarrer[3].NoFault := FALSE;
   MouldCarrer[3].MachineAutomatic := FALSE;
   MouldCarrer[3].MHAutomatic := FALSE;
   MouldCarrer[3].RobotAutomatic := FALSE;
   MouldCarrer[3].WetShot := FALSE;
   MouldCarrer[3].CycleRun := FALSE;
   MouldCarrer[3].ReadyForShot := FALSE;
   MouldCarrer[3].ShotRun := FALSE;
   MouldCarrer[3].CPsisForward := FALSE;
   MouldCarrer[3].Status_Spare_01 := FALSE;
   MouldCarrer[3].Status_Spare_02 := FALSE;
   MouldCarrer[3].Status_Spare_03 := FALSE;
   MouldCarrer[3].Status_Spare_04 := FALSE;
   MouldCarrer[3].Status_Spare_05 := FALSE;
   MouldCarrer[3].Status_Spare_06 := FALSE;
   MouldCarrer[3].Status_Spare_07 := FALSE;
   MouldCarrer[3].ProgNumber := FALSE;
   MouldCarrer[3].Fault_01 := FALSE;
   MouldCarrer[3].Fault_02 := FALSE;
   MouldCarrer[3].Fault_03 := FALSE;
   MouldCarrer[3].Fault_04 := FALSE;
   MouldCarrer[3].Fault_05 := FALSE;
   MouldCarrer[3].Fault_06 := FALSE;
   MouldCarrer[3].Fault_07 := FALSE;
   MouldCarrer[3].Fault_08 := FALSE;
   MouldCarrer[4].Preparation := FALSE;
   MouldCarrer[4].StartFoaming := FALSE;
   MouldCarrer[4].IN_Spare_01 := FALSE;
   MouldCarrer[4].IN_Spare_02 := FALSE;
   MouldCarrer[4].IN_Spare_03 := FALSE;
   MouldCarrer[4].IN_Spare_04 := FALSE;
   MouldCarrer[4].IN_Spare_05 := FALSE;
   MouldCarrer[4].IN_Spare_06 := FALSE;
   MouldCarrer[4].ShotEnds := FALSE;
   MouldCarrer[4].Break := FALSE;
   MouldCarrer[4].OUT_Spare_01 := FALSE;
   MouldCarrer[4].OUT_Spare_02 := FALSE;
   MouldCarrer[4].OUT_Spare_03 := FALSE;
   MouldCarrer[4].OUT_Spare_04 := FALSE;
   MouldCarrer[4].OUT_Spare_05 := FALSE;
   MouldCarrer[4].OUT_Spare_06 := FALSE;
   MouldCarrer[4].NoFault := FALSE;
   // 983 more start values not shown
END_DATA_BLOCK

DATA_BLOCK "DB122_FlowIndexState"   // DB122
TITLE = Flow-Index and Flow-State of modul-channel
{ S7_Optimized_Access := 'FALSE' }
AUTHOR : KT242
NAME : Flow
VERSION : 0.1
   VAR
      MeteringUnit : Array[0..12] of "UDT121_DF_Chanel";
   END_VAR
BEGIN
   MeteringUnit[0].OUT_PROCAN.FlowIndex.FlowIndex0 := FALSE;
   MeteringUnit[0].OUT_PROCAN.FlowIndex.FlowIndex1 := FALSE;
   MeteringUnit[0].OUT_PROCAN.FlowIndex.FlowIndex2 := FALSE;
   MeteringUnit[0].OUT_PROCAN.FlowIndex.FlowIndex3 := FALSE;
   MeteringUnit[0].OUT_PROCAN.FlowIndex.Spare4 := FALSE;
   MeteringUnit[0].OUT_PROCAN.FlowIndex.Notclosedloop := FALSE;
   MeteringUnit[0].OUT_PROCAN.FlowIndex.StartQPB := FALSE;
   MeteringUnit[0].OUT_PROCAN.FlowIndex.Enableclosedloop := FALSE;
   MeteringUnit[0].OUT_PROCAN.TandemComand := 16#0000;
   MeteringUnit[0].OUT_PROCAN.SpareWord := 16#0000;
   MeteringUnit[0].OUT_PROCAN.Spare_DWORD_56 := 16#0000_0000;
   MeteringUnit[0].IN_PROCAN.Flowrate := 0;
   MeteringUnit[0].IN_PROCAN.PistonPosition := 0;
   MeteringUnit[0].IN_PROCAN.TandemStatus := 16#0000;
   MeteringUnit[0].IN_PROCAN.Spare_DWORD_96 := 16#0000_0000;
   MeteringUnit[1].OUT_PROCAN.FlowIndex.FlowIndex0 := FALSE;
   MeteringUnit[1].OUT_PROCAN.FlowIndex.FlowIndex1 := FALSE;
   MeteringUnit[1].OUT_PROCAN.FlowIndex.FlowIndex2 := FALSE;
   MeteringUnit[1].OUT_PROCAN.FlowIndex.FlowIndex3 := FALSE;
   MeteringUnit[1].OUT_PROCAN.FlowIndex.Spare4 := FALSE;
   MeteringUnit[1].OUT_PROCAN.FlowIndex.Notclosedloop := FALSE;
   MeteringUnit[1].OUT_PROCAN.FlowIndex.StartQPB := FALSE;
   MeteringUnit[1].OUT_PROCAN.FlowIndex.Enableclosedloop := FALSE;
   MeteringUnit[1].OUT_PROCAN.TandemComand := 16#0000;
   MeteringUnit[1].OUT_PROCAN.SpareWord := 16#0000;
   MeteringUnit[1].OUT_PROCAN.Spare_DWORD_56 := 16#0000_0000;
   MeteringUnit[1].IN_PROCAN.Flowrate := 0;
   MeteringUnit[1].IN_PROCAN.PistonPosition := 0;
   MeteringUnit[1].IN_PROCAN.TandemStatus := 16#0000;
   MeteringUnit[1].IN_PROCAN.Spare_DWORD_96 := 16#0000_0000;
   MeteringUnit[2].OUT_PROCAN.FlowIndex.FlowIndex0 := FALSE;
   MeteringUnit[2].OUT_PROCAN.FlowIndex.FlowIndex1 := FALSE;
   MeteringUnit[2].OUT_PROCAN.FlowIndex.FlowIndex2 := FALSE;
   MeteringUnit[2].OUT_PROCAN.FlowIndex.FlowIndex3 := FALSE;
   MeteringUnit[2].OUT_PROCAN.FlowIndex.Spare4 := FALSE;
   MeteringUnit[2].OUT_PROCAN.FlowIndex.Notclosedloop := FALSE;
   MeteringUnit[2].OUT_PROCAN.FlowIndex.StartQPB := FALSE;
   MeteringUnit[2].OUT_PROCAN.FlowIndex.Enableclosedloop := FALSE;
   MeteringUnit[2].OUT_PROCAN.TandemComand := 16#0000;
   MeteringUnit[2].OUT_PROCAN.SpareWord := 16#0000;
   MeteringUnit[2].OUT_PROCAN.Spare_DWORD_56 := 16#0000_0000;
   MeteringUnit[2].IN_PROCAN.Flowrate := 0;
   MeteringUnit[2].IN_PROCAN.PistonPosition := 0;
   MeteringUnit[2].IN_PROCAN.TandemStatus := 16#0000;
   MeteringUnit[2].IN_PROCAN.Spare_DWORD_96 := 16#0000_0000;
   MeteringUnit[3].OUT_PROCAN.FlowIndex.FlowIndex0 := FALSE;
   MeteringUnit[3].OUT_PROCAN.FlowIndex.FlowIndex1 := FALSE;
   MeteringUnit[3].OUT_PROCAN.FlowIndex.FlowIndex2 := FALSE;
   MeteringUnit[3].OUT_PROCAN.FlowIndex.FlowIndex3 := FALSE;
   MeteringUnit[3].OUT_PROCAN.FlowIndex.Spare4 := FALSE;
   MeteringUnit[3].OUT_PROCAN.FlowIndex.Notclosedloop := FALSE;
   MeteringUnit[3].OUT_PROCAN.FlowIndex.StartQPB := FALSE;
   MeteringUnit[3].OUT_PROCAN.FlowIndex.Enableclosedloop := FALSE;
   MeteringUnit[3].OUT_PROCAN.TandemComand := 16#0000;
   MeteringUnit[3].OUT_PROCAN.SpareWord := 16#0000;
   MeteringUnit[3].OUT_PROCAN.Spare_DWORD_56 := 16#0000_0000;
   MeteringUnit[3].IN_PROCAN.Flowrate := 0;
   MeteringUnit[3].IN_PROCAN.PistonPosition := 0;
   MeteringUnit[3].IN_PROCAN.TandemStatus := 16#0000;
   MeteringUnit[3].IN_PROCAN.Spare_DWORD_96 := 16#0000_0000;
   MeteringUnit[4].OUT_PROCAN.FlowIndex.FlowIndex0 := FALSE;
   MeteringUnit[4].OUT_PROCAN.FlowIndex.FlowIndex1 := FALSE;
   MeteringUnit[4].OUT_PROCAN.FlowIndex.FlowIndex2 := FALSE;
   MeteringUnit[4].OUT_PROCAN.FlowIndex.FlowIndex3 := FALSE;
   MeteringUnit[4].OUT_PROCAN.FlowIndex.Spare4 := FALSE;
   MeteringUnit[4].OUT_PROCAN.FlowIndex.Notclosedloop := FALSE;
   MeteringUnit[4].OUT_PROCAN.FlowIndex.StartQPB := FALSE;
   MeteringUnit[4].OUT_PROCAN.FlowIndex.Enableclosedloop := FALSE;
   MeteringUnit[4].OUT_PROCAN.TandemComand := 16#0000;
   MeteringUnit[4].OUT_PROCAN.SpareWord := 16#0000;
   MeteringUnit[4].OUT_PROCAN.Spare_DWORD_56 := 16#0000_0000;
   MeteringUnit[4].IN_PROCAN.Flowrate := 0;
   MeteringUnit[4].IN_PROCAN.PistonPosition := 0;
   MeteringUnit[4].IN_PROCAN.TandemStatus := 16#0000;
   MeteringUnit[4].IN_PROCAN.Spare_DWORD_96 := 16#0000_0000;
   MeteringUnit[5].OUT_PROCAN.FlowIndex.FlowIndex0 := FALSE;
   MeteringUnit[5].OUT_PROCAN.FlowIndex.FlowIndex1 := FALSE;
   MeteringUnit[5].OUT_PROCAN.FlowIndex.FlowIndex2 := FALSE;
   MeteringUnit[5].OUT_PROCAN.FlowIndex.FlowIndex3 := FALSE;
   MeteringUnit[5].OUT_PROCAN.FlowIndex.Spare4 := FALSE;
   MeteringUnit[5].OUT_PROCAN.FlowIndex.Notclosedloop := FALSE;
   MeteringUnit[5].OUT_PROCAN.FlowIndex.StartQPB := FALSE;
   MeteringUnit[5].OUT_PROCAN.FlowIndex.Enableclosedloop := FALSE;
   MeteringUnit[5].OUT_PROCAN.TandemComand := 16#0000;
   MeteringUnit[5].OUT_PROCAN.SpareWord := 16#0000;
   MeteringUnit[5].OUT_PROCAN.Spare_DWORD_56 := 16#0000_0000;
   MeteringUnit[5].IN_PROCAN.Flowrate := 0;
   MeteringUnit[5].IN_PROCAN.PistonPosition := 0;
   MeteringUnit[5].IN_PROCAN.TandemStatus := 16#0000;
   MeteringUnit[5].IN_PROCAN.Spare_DWORD_96 := 16#0000_0000;
   MeteringUnit[6].OUT_PROCAN.FlowIndex.FlowIndex0 := FALSE;
   MeteringUnit[6].OUT_PROCAN.FlowIndex.FlowIndex1 := FALSE;
   MeteringUnit[6].OUT_PROCAN.FlowIndex.FlowIndex2 := FALSE;
   MeteringUnit[6].OUT_PROCAN.FlowIndex.FlowIndex3 := FALSE;
   MeteringUnit[6].OUT_PROCAN.FlowIndex.Spare4 := FALSE;
   MeteringUnit[6].OUT_PROCAN.FlowIndex.Notclosedloop := FALSE;
   MeteringUnit[6].OUT_PROCAN.FlowIndex.StartQPB := FALSE;
   MeteringUnit[6].OUT_PROCAN.FlowIndex.Enableclosedloop := FALSE;
   MeteringUnit[6].OUT_PROCAN.TandemComand := 16#0000;
   MeteringUnit[6].OUT_PROCAN.SpareWord := 16#0000;
   MeteringUnit[6].OUT_PROCAN.Spare_DWORD_56 := 16#0000_0000;
   MeteringUnit[6].IN_PROCAN.Flowrate := 0;
   MeteringUnit[6].IN_PROCAN.PistonPosition := 0;
   MeteringUnit[6].IN_PROCAN.TandemStatus := 16#0000;
   MeteringUnit[6].IN_PROCAN.Spare_DWORD_96 := 16#0000_0000;
   MeteringUnit[7].OUT_PROCAN.FlowIndex.FlowIndex0 := FALSE;
   MeteringUnit[7].OUT_PROCAN.FlowIndex.FlowIndex1 := FALSE;
   MeteringUnit[7].OUT_PROCAN.FlowIndex.FlowIndex2 := FALSE;
   MeteringUnit[7].OUT_PROCAN.FlowIndex.FlowIndex3 := FALSE;
   MeteringUnit[7].OUT_PROCAN.FlowIndex.Spare4 := FALSE;
   MeteringUnit[7].OUT_PROCAN.FlowIndex.Notclosedloop := FALSE;
   MeteringUnit[7].OUT_PROCAN.FlowIndex.StartQPB := FALSE;
   MeteringUnit[7].OUT_PROCAN.FlowIndex.Enableclosedloop := FALSE;
   MeteringUnit[7].OUT_PROCAN.TandemComand := 16#0000;
   MeteringUnit[7].OUT_PROCAN.SpareWord := 16#0000;
   MeteringUnit[7].OUT_PROCAN.Spare_DWORD_56 := 16#0000_0000;
   MeteringUnit[7].IN_PROCAN.Flowrate := 0;
   MeteringUnit[7].IN_PROCAN.PistonPosition := 0;
   MeteringUnit[7].IN_PROCAN.TandemStatus := 16#0000;
   MeteringUnit[7].IN_PROCAN.Spare_DWORD_96 := 16#0000_0000;
   MeteringUnit[8].OUT_PROCAN.FlowIndex.FlowIndex0 := FALSE;
   MeteringUnit[8].OUT_PROCAN.FlowIndex.FlowIndex1 := FALSE;
   MeteringUnit[8].OUT_PROCAN.FlowIndex.FlowIndex2 := FALSE;
   MeteringUnit[8].OUT_PROCAN.FlowIndex.FlowIndex3 := FALSE;
   MeteringUnit[8].OUT_PROCAN.FlowIndex.Spare4 := FALSE;
   MeteringUnit[8].OUT_PROCAN.FlowIndex.Notclosedloop := FALSE;
   MeteringUnit[8].OUT_PROCAN.FlowIndex.StartQPB := FALSE;
   MeteringUnit[8].OUT_PROCAN.FlowIndex.Enableclosedloop := FALSE;
   MeteringUnit[8].OUT_PROCAN.TandemComand := 16#0000;
   MeteringUnit[8].OUT_PROCAN.SpareWord := 16#0000;
   MeteringUnit[8].OUT_PROCAN.Spare_DWORD_56 := 16#0000_0000;
   MeteringUnit[8].IN_PROCAN.Flowrate := 0;
   MeteringUnit[8].IN_PROCAN.PistonPosition := 0;
   MeteringUnit[8].IN_PROCAN.TandemStatus := 16#0000;
   MeteringUnit[8].IN_PROCAN.Spare_DWORD_96 := 16#0000_0000;
   MeteringUnit[9].OUT_PROCAN.FlowIndex.FlowIndex0 := FALSE;
   MeteringUnit[9].OUT_PROCAN.FlowIndex.FlowIndex1 := FALSE;
   MeteringUnit[9].OUT_PROCAN.FlowIndex.FlowIndex2 := FALSE;
   MeteringUnit[9].OUT_PROCAN.FlowIndex.FlowIndex3 := FALSE;
   MeteringUnit[9].OUT_PROCAN.FlowIndex.Spare4 := FALSE;
   MeteringUnit[9].OUT_PROCAN.FlowIndex.Notclosedloop := FALSE;
   MeteringUnit[9].OUT_PROCAN.FlowIndex.StartQPB := FALSE;
   MeteringUnit[9].OUT_PROCAN.FlowIndex.Enableclosedloop := FALSE;
   MeteringUnit[9].OUT_PROCAN.TandemComand := 16#0000;
   MeteringUnit[9].OUT_PROCAN.SpareWord := 16#0000;
   MeteringUnit[9].OUT_PROCAN.Spare_DWORD_56 := 16#0000_0000;
   MeteringUnit[9].IN_PROCAN.Flowrate := 0;
   MeteringUnit[9].IN_PROCAN.PistonPosition := 0;
   MeteringUnit[9].IN_PROCAN.TandemStatus := 16#0000;
   MeteringUnit[9].IN_PROCAN.Spare_DWORD_96 := 16#0000_0000;
   MeteringUnit[10].OUT_PROCAN.FlowIndex.FlowIndex0 := FALSE;
   MeteringUnit[10].OUT_PROCAN.FlowIndex.FlowIndex1 := FALSE;
   MeteringUnit[10].OUT_PROCAN.FlowIndex.FlowIndex2 := FALSE;
   MeteringUnit[10].OUT_PROCAN.FlowIndex.FlowIndex3 := FALSE;
   MeteringUnit[10].OUT_PROCAN.FlowIndex.Spare4 := FALSE;
   MeteringUnit[10].OUT_PROCAN.FlowIndex.Notclosedloop := FALSE;
   MeteringUnit[10].OUT_PROCAN.FlowIndex.StartQPB := FALSE;
   MeteringUnit[10].OUT_PROCAN.FlowIndex.Enableclosedloop := FALSE;
   MeteringUnit[10].OUT_PROCAN.TandemComand := 16#0000;
   MeteringUnit[10].OUT_PROCAN.SpareWord := 16#0000;
   MeteringUnit[10].OUT_PROCAN.Spare_DWORD_56 := 16#0000_0000;
   MeteringUnit[10].IN_PROCAN.Flowrate := 0;
   MeteringUnit[10].IN_PROCAN.PistonPosition := 0;
   MeteringUnit[10].IN_PROCAN.TandemStatus := 16#0000;
   MeteringUnit[10].IN_PROCAN.Spare_DWORD_96 := 16#0000_0000;
   MeteringUnit[11].OUT_PROCAN.FlowIndex.FlowIndex0 := FALSE;
   MeteringUnit[11].OUT_PROCAN.FlowIndex.FlowIndex1 := FALSE;
   MeteringUnit[11].OUT_PROCAN.FlowIndex.FlowIndex2 := FALSE;
   MeteringUnit[11].OUT_PROCAN.FlowIndex.FlowIndex3 := FALSE;
   MeteringUnit[11].OUT_PROCAN.FlowIndex.Spare4 := FALSE;
   MeteringUnit[11].OUT_PROCAN.FlowIndex.Notclosedloop := FALSE;
   MeteringUnit[11].OUT_PROCAN.FlowIndex.StartQPB := FALSE;
   MeteringUnit[11].OUT_PROCAN.FlowIndex.Enableclosedloop := FALSE;
   MeteringUnit[11].OUT_PROCAN.TandemComand := 16#0000;
   MeteringUnit[11].OUT_PROCAN.SpareWord := 16#0000;
   MeteringUnit[11].OUT_PROCAN.Spare_DWORD_56 := 16#0000_0000;
   MeteringUnit[11].IN_PROCAN.Flowrate := 0;
   MeteringUnit[11].IN_PROCAN.PistonPosition := 0;
   MeteringUnit[11].IN_PROCAN.TandemStatus := 16#0000;
   MeteringUnit[11].IN_PROCAN.Spare_DWORD_96 := 16#0000_0000;
   MeteringUnit[12].OUT_PROCAN.FlowIndex.FlowIndex0 := FALSE;
   MeteringUnit[12].OUT_PROCAN.FlowIndex.FlowIndex1 := FALSE;
   MeteringUnit[12].OUT_PROCAN.FlowIndex.FlowIndex2 := FALSE;
   MeteringUnit[12].OUT_PROCAN.FlowIndex.FlowIndex3 := FALSE;
   MeteringUnit[12].OUT_PROCAN.FlowIndex.Spare4 := FALSE;
   MeteringUnit[12].OUT_PROCAN.FlowIndex.Notclosedloop := FALSE;
   MeteringUnit[12].OUT_PROCAN.FlowIndex.StartQPB := FALSE;
   MeteringUnit[12].OUT_PROCAN.FlowIndex.Enableclosedloop := FALSE;
   MeteringUnit[12].OUT_PROCAN.TandemComand := 16#0000;
   MeteringUnit[12].OUT_PROCAN.SpareWord := 16#0000;
   MeteringUnit[12].OUT_PROCAN.Spare_DWORD_56 := 16#0000_0000;
   MeteringUnit[12].IN_PROCAN.Flowrate := 0;
   MeteringUnit[12].IN_PROCAN.PistonPosition := 0;
   MeteringUnit[12].IN_PROCAN.TandemStatus := 16#0000;
   MeteringUnit[12].IN_PROCAN.Spare_DWORD_96 := 16#0000_0000;
END_DATA_BLOCK

DATA_BLOCK "DB123_MH_IO_Signals"   // DB123
TITLE = IO-Signals of mixinghead operation panel
{ S7_Optimized_Access := 'FALSE' }
AUTHOR : KT242
NAME : MHead
VERSION : 0.1
   VAR
      MH : Array[0..16] of "UDT123_MH_Chanel";
   END_VAR
BEGIN
END_DATA_BLOCK

